               ELSIF (#statCountChannelPos = #CONST_CHANNEL_POS1)
               THEN
                   #statCurrentPos2 := #statCountChannelPos;
                   #statTimeImpulseSave2 := #statDeltaTimeImpulse;
                   #statTimePauseSave2 := #statDeltaTimePause;
                   #statTimeToImpulse := #statTimeToImpulse + #statDeltaTimeImpulse + #statDeltaTimePause;

                   IF ((#statDeltaTimePause >= #TIME_PAUSE1_MIN)
                       AND (#statDeltaTimePause <= #TIME_PAUSE1_MAX))
                   THEN
                       #statChannelActive2 := true;
                       #statCountChannelPos := #CONST_CHANNEL_POS2; // go to next pos 2
                   END_IF;

                   IF ((#statDeltaTimePause >= #TIME_PAUSE2_MIN)
                       AND (#statDeltaTimePause <= #TIME_PAUSE2_MAX))
                   THEN
                       #statChannelActive2 := false;
                       #statChannelActive3 := true;
                       #statCountChannelPos := #CONST_CHANNEL_POS2; // go to next Pos 2
                   END_IF;

                   IF ((#statDeltaTimePause >= #TIME_PAUSE3_MIN)
                       AND (#statDeltaTimePause <= #TIME_PAUSE3_MAX))
                   THEN
                       #statChannelActive2 := false;
                       #statChannelActive3 := false;
                       #statChannelActive4 := true;
                       #statCountChannelPos := #CONST_INT_0;
                   END_IF;

               ELSIF (#statCountChannelPos = #CONST_CHANNEL_POS2)
               THEN
                   #statCurrentPos3 := #statCountChannelPos;
                   #statTimeImpulseSave3 := #statDeltaTimeImpulse;
                   #statTimePauseSave3 := #statDeltaTimePause;
                   #statTimeToImpulse := #statTimeToImpulse + #statDeltaTimeImpulse + #statDeltaTimePause;

                   IF ((#statDeltaTimePause >= #TIME_PAUSE1_MIN)
                       AND (#statDeltaTimePause <= #TIME_PAUSE1_MAX))
                   THEN
                       #statChannelActive3 := true;
                       #statCountChannelPos := #CONST_CHANNEL_POS3; // go to next pos 3
                   END_IF;

                   IF ((#statDeltaTimePause >= #TIME_PAUSE2_MIN)
                       AND (#statDeltaTimePause <= #TIME_PAUSE2_MAX))
                   THEN
                       #statChannelActive3 := false;
                       #statChannelActive4 := true;
                       #statCountChannelPos := #CONST_INT_0;
                   END_IF;

               ELSIF (#statCountChannelPos = #CONST_CHANNEL_POS3)
               THEN
                   #statCurrentPos4 := #statCountChannelPos;
                   #statTimeImpulseSave4 := #statDeltaTimeImpulse;
                   #statTimePauseSave4 := #statDeltaTimePause;
                   #statTimeToImpulse := #statTimeToImpulse + #statDeltaTimeImpulse + #statDeltaTimePause;

                   IF ((#statDeltaTimePause >= #TIME_PAUSE1_MIN)
                       AND (#statDeltaTimePause <= #TIME_PAUSE1_MAX))
                   THEN
                       #statChannelActive4 := true;
                   END_IF;
                   #statCountChannelPos := #CONST_INT_0; // go to pos 0
               END_IF;
           END_IF;

       #STATE_ERROR:
           #error := true;
           #busy := false;
           #done := false;
           #statSysTimerStart := false;
           #statWatchDogTimerRisingStart := false;
           #statWatchDogTimerFallingStart := false;
           #status := #statStatus;
           #statStatus := #CONST_WORD_0;
           #statIndex := #STATE_IDLE;
       ELSE
           #statIndex := #STATE_IDLE;
   END_CASE;

   #instWatchDogTimerRising(IN := #statWatchDogTimerRisingStart,
                      PT := #CONST_WATCHDOG_TIMER,
                      Q=>#statWatchDogTimerRisingStop,
                      ET=>#statWatchDogTimerRisingRun);

   #instWatchDogTimerFalling(IN:=#statWatchDogTimerFallingStart,
                             PT:=#CONST_WATCHDOG_TIMER,
                             Q=>#statWatchDogTimerFallingStop,
                             ET=>#statWatchDogTimerFallingRun);


   #instSysTimer(IN:=#statSysTimerStart,
                 PT:=#CONST_CYCLETIME_TIMER,
                 Q=>#statSysTimerStop,
                 ET=>#statSysTimerRun);

   IF (#statWatchDogTimerRisingStop = TRUE)
       OR (#statWatchDogTimerFallingStop =true)
   THEN
       #statIndex := #STATE_ERROR;
       #statStatus := #CONST_ERROR_WATCHDOG_TIMER;
   END_IF;


   IF (#statSysTimerStop=true)
   THEN
       #statIndex := #STATE_ERROR;
       #statStatus := #CONST_ERROR_CYCLETIME_TIMER;
   END_IF;

   //Edge control
   #statImpulseOld := #impulse;
   #statResetOld := #reset;

   // Cycle time control
   #statSysTimeOld := #statSysTime;
END_FUNCTION_BLOCK

// ===== library types =====

TYPE "M_ZLT"
VERSION : 0.1
   STRUCT
      Fehl_empf : Bool;
      Fehl_Krit : Bool;
      Fehl_TO : Bool;
      STue_Abgl : Bool;
      Mel_Überlauf : Bool;
      Mel_Parameter : Bool;
      F_PW_Nr : Bool;
      Fehl_Senden : Bool;
      RM_ArbZeit : Bool;
      RM_Pause : Bool;
      RM_Schicht_1 : Bool;
      RM_Schicht_2 : Bool;
      RM_Schicht_3 : Bool;
      RM_Schicht_4 : Bool;
      RM_LSp : Bool;
      RM_Res : Bool;
   END_STRUCT;
END_TYPE

// folder: Audi_Bib/GF_Bausteine

FUNCTION_BLOCK "GF_GrFunktionen"   // FB200, SCL
{ S7_Optimized_Access := 'TRUE' }
VERSION : 0.1
   VAR_INPUT
      Quit_F : Bool;   // Quittierung Sicherheit/ Wiedereingliederung
      Init : Bool;
      TW_Res : Time;   // Zeitwert Resetzeit in 0,1s max 25sec
      TW_FQuit : Time;
   END_VAR
   VAR_OUTPUT
      F_Quit : Bool;
   END_VAR
   VAR
      R_TRIG_Instance : R_TRIG;
   END_VAR
   VAR RETAIN
      HMAnlauf : Bool;   // Hilfsmerker Anlauf
      HMAnl_ab : Bool;
      A_F_Quit : Bool;
      Quit_F_ab : Bool;
      Anl_Verzögerung : TON_TIME;
      IEC_Timer_0_Instance : TOF_TIME;
      Ret_SNC_RTCB : Int;
      Ret_WR_SYS : Int;
      T_Start_1 : Bool;
      T_abgel_1 : Bool;
      T_Start_2 : Bool;
      T_abgel_2 : Bool;
      Lfd_Nr_HText_1 : Int;
      Lfd_Nr_HText_2 : Int;
      "Tverz_Info-Text_1" : TON_TIME;
      "TVerz_Info-Text_2" : TON_TIME;
   END_VAR
   VAR_TEMP
      Stell_Zeit : DTL;
      S_1 : String;
      Ret_VAl : Int;
      T_Int : Int;
      UInt_1 : UInt;
      Zeit : String;
      Datum : String;
      X_Anzahl : Int;
      x : Int;
      Dat_Uhrz : String[24];
      HStr_3 : String[3];
   END_VAR
BEGIN
   (* Funktionsbeschreibung:                                                   Stand 6.5.2015
   ----------------------


   Baustein-Änderungen:
   --------------------
   Stand 9.6.2011  Identisch mit FB60 V 1.9 NSU Stand 18.2.2011
   Stand 22.9.2011  CPU-Meldungen aus Fehlermelde-OB´s angepasst (Adresse)
                    gemessene Zykluszeit "Mit" Rücksetzung eingefügt
   Stand 6.5.2015   Umstellung Takt-Merker auf Cyclic Interrupt-OB_s dadurch werden
                    keine CPU-Taktmerker mehr benötigt
   V0.1.7    Remanenz und Speicherreserve für Laden eingestellt



   *)                

   "VKE0":= false; "VS".VKE0 := false;                               // Vorbesetzung Systemmerker
   "VKE1":= true; "VS".VKE1 := true;
   "VS".Null := false;
   "VS".Eins := TRUE;
   "VS".Ohne := false;
   "VS".Mit := true;
   "VS".Mel_int := false;
   "VS".Kon_int := false;
   "VS".Sifa_int := false;

   "VS".Steu_ein := True;

   "VS".BliL := "VS"."Takt_0,5s";            // Blinktakte 500mSek
   "VS".BliS := "VS"."Takt_0,2s";              // Blinktakt 250mSek

   "VS"."ZTakt_0,1s" := false;                 // Zähltakt 100mSek.
   IF "VS"."Trig_0,1s" THEN
      "VS"."ZTakt_0,1s" := true;
      "VS"."Trig_0,1s" := false;
   END_IF;
   #R_TRIG_Instance(CLK:="VS"."Takt_0,5s", Q=>"VS".ZTakt_1s);               // Zähltakt 1Sekunde


   IF #HMAnlauf THEN #HMAnlauf:= false; "VS".Neustart:= false;  END_IF;       // Anlauf nach Neustart
   IF "VS".Neustart  THEN "VS".Anl_Verlae:= true; #HMAnlauf:= true; END_IF;
   #Anl_Verzögerung(IN:="VS".Anl_Verlae, PT:=#TW_Res,Q=>#HMAnl_ab );
   IF #HMAnl_ab THEN "VS".Anl_Verlae:= false; END_IF;
   "VS".Reset := "VS".Anl_Verlae;

   IF #HMAnl_ab OR "VS".Neustart  THEN #A_F_Quit:= true; END_IF;                        // F-Quit bilden
   #IEC_Timer_0_Instance(IN:=#A_F_Quit,  PT:=#TW_FQuit, Q=>#Quit_F_ab);
   IF #Quit_F_ab THEN #A_F_Quit:= false; END_IF;
   #F_Quit:= #A_F_Quit;

   // ************* Zykluszeit
   "GF_Zeitmessung"(Reset:="GF_Grund_DB".Res_Zeit[1],    // Zykluszeit errechnen
                    Mes_auswert:=true,
                    Zeit:="GF_Grund_DB".Zeit[1]);


   // CPU Zeit Stellen  Anstoss von Panel oder aus ZLT-Paket(Zeit-Synchronisation)
   IF "GF_Grund_DB".Stellbits.OP_Stell OR "GF_Grund_DB".Stellbits.Stell_ASCII THEN
      IF "GF_Grund_DB".Stellbits.Stell_ASCII THEN                                          // Zeitsynchronisation
         "GF_Grund_DB".Stellbits.Stell_ASCII := FALSE;                                                           //Stellzeit Typ DTL aus ASCII bilden
         Chars_TO_Strg(Chars := "GF_Grund_DB".Stell_Datum_Uhrzeit_ASCI.Jahr, pChars := 0, Cnt := 4,  Strg => #S_1);      //    Jahr
         #Stell_Zeit.YEAR := S_CONV(#S_1);
         Chars_TO_Strg(Chars := "GF_Grund_DB".Stell_Datum_Uhrzeit_ASCI.Monat, pChars := 0, Cnt := 2, Strg => #S_1);      //    Monat
         #Stell_Zeit.MONTH := S_CONV(#S_1);
         Chars_TO_Strg(Chars := "GF_Grund_DB".Stell_Datum_Uhrzeit_ASCI.Tag, pChars := 0, Cnt := 2, Strg => #S_1);        //    Tag
         #Stell_Zeit.DAY := S_CONV(#S_1);

         Chars_TO_Strg(Chars := "GF_Grund_DB".Stell_Datum_Uhrzeit_ASCI.Stunde, pChars := 0, Cnt := 2, Strg => #S_1);     //    Stunde
         #Stell_Zeit.HOUR := S_CONV(#S_1);
         Chars_TO_Strg(Chars := "GF_Grund_DB".Stell_Datum_Uhrzeit_ASCI.Minute, pChars := 0, Cnt := 2, Strg => #S_1);     //    Minute
         #Stell_Zeit.MINUTE := S_CONV(#S_1);
         Chars_TO_Strg(Chars := "GF_Grund_DB".Stell_Datum_Uhrzeit_ASCI.Sekunde, pChars := 0, Cnt := 2, Strg => #S_1);    //    Sekunde
         #Stell_Zeit.SECOND := S_CONV(#S_1);

         Chars_TO_Strg(Chars := "GF_Grund_DB".Stell_Datum_Uhrzeit_ASCI.MilliSek, pChars := 0, Cnt := 3, Strg => #S_1);   //    Millisekunde
         #Stell_Zeit.NANOSECOND := S_CONV(#S_1);
         #S_1 := S_CONV("GF_Grund_DB".Stell_Datum_Uhrzeit_ASCI.Wochentag);                                       //    Wochentag
         #Stell_Zeit.WEEKDAY := S_CONV(#S_1);

         "GF_Grund_DB".Stell_Datum_Uhrzeit := #Stell_Zeit;
         END_IF;

      IF "GF_Grund_DB".Stellbits.OP_Stell THEN                                 // Uhrzeit stellen von TP (Format DTL)
         "GF_Grund_DB".Stellbits.OP_Stell := false;
         #Stell_Zeit := "GF_Grund_DB".Stell_Datum_Uhrzeit;
      END_IF;

      #Ret_WR_SYS := WR_SYS_T(#Stell_Zeit);           // Uhrzeit stellen
      "GF_Grund_DB".Ret_Val := #Ret_VAl;

      #Ret_SNC_RTCB := SNC_RTCB();                      // Zeitsynchronisation nachtriggern
   END_IF;
   #T_Int := #Ret_SNC_RTCB; #T_Int := #Ret_WR_SYS;


   // ******************* CPU-Zeit auslesen
   //  Datum
   #Ret_VAl:=RD_LOC_T("GF_Grund_DB".Akt_Datum_Uhrzeit);                                                           // Aktuelle Datum/Zeit im Format DTL
   #S_1:=S_CONV("GF_Grund_DB".Akt_Datum_Uhrzeit.YEAR);                                                      // Umsetzung DTL in ASCII  Jahr
   #S_1:=RIGHT(IN:=#S_1, L:=4);
   #UInt_1 := 4;
   Strg_TO_Chars(Strg:=#S_1, pChars:=0,Cnt=>#UInt_1 , Chars:="GF_Grund_DB".Akt_Datum_Uhrzeit_ASCII.Datum.Jahr);
   #Datum := #S_1;
   #S_1:=S_CONV("GF_Grund_DB".Akt_Datum_Uhrzeit.MONTH);                                                     // Monat 
   #S_1 := REPLACE(IN1 := #S_1, IN2 := '0', L := 1, P := 1);
   #S_1:=RIGHT(IN:=#S_1, L:=2);
   Strg_TO_Chars(Strg:=#S_1, pChars:=0,Cnt=>#UInt_1, Chars:="GF_Grund_DB".Akt_Datum_Uhrzeit_ASCII.Datum.Monat);
   #Datum :=CONCAT(IN1:=#Datum, IN2:=#S_1);
   #S_1:=S_CONV("GF_Grund_DB".Akt_Datum_Uhrzeit.DAY);                                                       // Tag
   #S_1 := REPLACE(IN1 := #S_1, IN2 := '0', L := 1, P := 1);
   #S_1 := RIGHT(IN := #S_1, L := 2);
   Strg_TO_Chars(Strg:=#S_1, pChars:=0,Cnt=>#UInt_1, Chars:="GF_Grund_DB".Akt_Datum_Uhrzeit_ASCII.Datum.Tag);
   "GF_Grund_DB".Akt_Datum_Uhrzeit_ASCII.Datum.YYYYMMDD := CONCAT(IN1 := #Datum, IN2 := #S_1);

   // ***************** Zeit
   #S_1:=S_CONV("GF_Grund_DB".Akt_Datum_Uhrzeit.HOUR);                                                       // Stunde
   #S_1 := REPLACE(IN1 := #S_1, IN2 := '0', L := 1, P := 1);
   #S_1 := RIGHT(IN := #S_1, L := 2);
   Strg_TO_Chars(Strg:=#S_1, pChars:=0,Cnt=>#UInt_1, Chars:="GF_Grund_DB".Akt_Datum_Uhrzeit_ASCII.Zeit.Stunde);
   #Zeit := #S_1;
   #S_1:=S_CONV("GF_Grund_DB".Akt_Datum_Uhrzeit.MINUTE);                                                    // Minute
   #S_1 := REPLACE(IN1 := #S_1, IN2 := '0', L := 1, P := 1);
   #S_1:=RIGHT(IN:=#S_1, L:=2);
   Strg_TO_Chars(Strg:=#S_1, pChars:=0,Cnt=>#UInt_1, Chars:="GF_Grund_DB".Akt_Datum_Uhrzeit_ASCII.Zeit.Minute);
   #Zeit := CONCAT(IN1 := #Zeit, IN2 := #S_1); 
   #S_1:=S_CONV("GF_Grund_DB".Akt_Datum_Uhrzeit.SECOND);                                                    // Sekunde
   #S_1 := REPLACE(IN1 := #S_1, IN2 := '0', L := 1, P := 1);
   #S_1:=RIGHT(IN:=#S_1, L:=2);
   Strg_TO_Chars(Strg:=#S_1, pChars:=0,Cnt=>#UInt_1, Chars:="GF_Grund_DB".Akt_Datum_Uhrzeit_ASCII.Zeit.Sekunde);
   "GF_Grund_DB".Akt_Datum_Uhrzeit_ASCII.Zeit.HHMMSS := CONCAT(IN1 := #Zeit, IN2 := #S_1);

   #S_1:=S_CONV("GF_Grund_DB".Akt_Datum_Uhrzeit.NANOSECOND);                                                                                                                        
   // Milli-Sekunde
   #S_1:=MID(IN:=#S_1, L:=3, P:=3);
   Strg_TO_Chars(Strg:=#S_1, pChars:=0,Cnt=>#UInt_1, Chars:="GF_Grund_DB".Akt_Datum_Uhrzeit_ASCII.Zeit.MilliSek);
   #S_1:=S_CONV("GF_Grund_DB".Akt_Datum_Uhrzeit.WEEKDAY);                                                   // Wochentag
   #S_1:=RIGHT(IN:=#S_1, L:=1);
   "GF_Grund_DB".Akt_Datum_Uhrzeit_ASCII.Wochentag :=S_CONV(#S_1);

   //*********** Zeitformat für MA-PC (Fuchs-Paket) bereitstellen
   #Dat_Uhrz := "GF_Grund_DB".Akt_Datum_Uhrzeit_ASCII.Datum.YYYYMMDD;
   #Dat_Uhrz := INSERT(IN1 := #Dat_Uhrz, IN2 := '-', P := 4);                                          // YYYY-MMTT
   #Dat_Uhrz := INSERT(IN1 := #Dat_Uhrz, IN2 := '-', P := 7);                                          // YYYY-MM-TT
   #Dat_Uhrz := INSERT(IN1 := #Dat_Uhrz, IN2 := '  ', P := 11);                                        // YYYY-MM-TT__
   #Dat_Uhrz := INSERT(IN1 := #Dat_Uhrz, IN2 := "GF_Grund_DB".Akt_Datum_Uhrzeit_ASCII.Zeit.HHMMSS, P := 12);   // 
   #Dat_Uhrz := INSERT(IN1 := #Dat_Uhrz, IN2 := ':', P := 14);                                         // YYYY-MM-TT__hh:mmss
   #Dat_Uhrz := INSERT(IN1 := #Dat_Uhrz, IN2 := ':', P := 17);                                         // YYYY-MM-TT__hh:mm:ss
   #Dat_Uhrz := INSERT(IN1 := #Dat_Uhrz, IN2 := ':', P := 20);                                         // YYYY-MM-TT__hh:mm:ss:
   Chars_TO_Strg(Chars := "GF_Grund_DB".Akt_Datum_Uhrzeit_ASCII.Zeit.MilliSek,
                 pChars := 0, Cnt := 3,Strg => #HStr_3);
   #Dat_Uhrz := INSERT(IN1 := #Dat_Uhrz, IN2 := #HStr_3, P := 21);                                     // YYYY-MM-TT__hh:mm:ss:mmm
   "GF_Grund_DB".Zeit_Ma_PC := #Dat_Uhrz;

   // *********  globale Visu Info-Texte nach 5 Sek freigaben
   IF "GF_Visu_allg".H_Text_1."umlfd.Nr" <> #Lfd_Nr_HText_1 AND "GF_Visu_allg".H_Text_1.Pult <> 'X'  THEN
      #Lfd_Nr_HText_1 := "GF_Visu_allg".H_Text_1."umlfd.Nr";
      #T_Start_1 := true;
   END_IF;
   #"Tverz_Info-Text_1"(IN := #T_Start_1, PT := T#5s, Q => #T_abgel_1);
   IF #T_abgel_1 THEN
      "GF_Visu_allg".H_Text_1."umlfd.Nr" := 0;
      "GF_Visu_allg".H_Text_1.Pult := 'X';
      "GF_Visu_allg".H_Text_1.Stellglied := ' ';
      "GF_Visu_allg".H_Text_1.H_Text := ' ';
      #T_Start_1 := false;
   END_IF;

   IF "GF_Visu_allg".H_Text_2."umlfd.Nr" <> #Lfd_Nr_HText_2 AND "GF_Visu_allg".H_Text_2.Pult <> 'X' THEN
      #Lfd_Nr_HText_2 := "GF_Visu_allg".H_Text_2."umlfd.Nr";
      #T_Start_2 := true;
   END_IF;
   #"TVerz_Info-Text_2"(IN := #T_Start_2, PT := T#5s, Q => #T_abgel_2);
   IF #T_abgel_2 THEN
      "GF_Visu_allg".H_Text_2."umlfd.Nr" := 0;
      "GF_Visu_allg".H_Text_2.Pult := 'X';
      "GF_Visu_allg".H_Text_2.Stellglied := ' ';
      "GF_Visu_allg".H_Text_2.H_Text := ' ';
      #T_Start_2 := false;
   END_IF;

   // ***********************  Initialisierungen
   IF #Init OR "VS".Neustart THEN
      #T_Start_1 := false;   #T_abgel_1 := false;
      #T_Start_2 := false;   #T_abgel_2 := false;

      "GF_Visu_allg".H_Text_1.Pult := 'X';
      "GF_Visu_allg".H_Text_1."umlfd.Nr" := 0;
      "GF_Visu_allg".H_Text_2.Pult := 'X';
      "GF_Visu_allg".H_Text_2."umlfd.Nr" := 0;

       #X_Anzahl := "GF_An_Vor_St".max_Anzahl;                         // An/Vorwahlen
       FOR #x := 1 TO #X_Anzahl DO                                     //   Eintrag Array-NR. in Array-Element NR
           "GF_An_Vor_St".An_Vorw[#x].AnVisu.Nr := #x;
           "GF_An_Vor_St".An_Vorw[#x].AnVisu.Bed_Station := 'xxxx';
           "GF_An_Vor_St".An_Vorw[#x].AnVisu.Bezeichnung := '    ';
           "GF_An_Vor_St".An_Vorw[#x].AnVisu.Status := 0;
       END_FOR;

       #X_Anzahl := "GF_LastSp_St".max_Anzahl;                         // Lastspannungen
       FOR #x := 1 TO #X_Anzahl DO                                     // Eintrag Array-NR. in Array-Element NR
           "GF_LastSp_St".LastSp[#x].AnVisu.Nr := #x;
           "GF_LastSp_St".LastSp[#x].AnVisu.Bed_Station := 'xxxx';
           "GF_LastSp_St".LastSp[#x].AnVisu.Bezeichnung := '    ';
           "GF_LastSp_St".LastSp[#x].AnVisu.Status := 0;
       END_FOR;

       #X_Anzahl := "GF_BetrArt_St".max_Anzahl;                        // Betriebsarten
       FOR #x := 1 TO #X_Anzahl DO                                     // Eintrag Array-NR. in Array-Element NR
           "GF_BetrArt_St".BetrArt[#x].AnVisu.Nr := #x;
           "GF_BetrArt_St".BetrArt[#x].AnVisu.Bed_Station := 'xxxx';
           "GF_BetrArt_St".BetrArt[#x].AnVisu.Bezeichnung := '    ';
           "GF_BetrArt_St".BetrArt[#x].AnVisu.Status := 0;
       END_FOR;

       #X_Anzahl := "GF_HBed_Obj_St".max_Anzahl;                       // Hand-Bedien-Objekte
       FOR #x := 1 TO #X_Anzahl DO                                     // Eintrag Array-NR. in Array-Element NR
           "GF_HBed_Obj_St".Modul[#x].Nr := #x;
       END_FOR;

       #X_Anzahl := 8;                                                 // Meldekanäle initialisieren
       FOR #x := 1 TO #X_Anzahl DO                                 
           "GF_Visu_allg".SS.Kanal[#x].Belegung.Pult_Name := 'xxxx';
       END_FOR;
   END_IF;
END_FUNCTION_BLOCK

FUNCTION "GF_Zeitmessung" : Void   // FC205, SCL
{ S7_Optimized_Access := 'TRUE' }
VERSION : 0.1
   VAR_INPUT
      Reset : Bool;   // Reset gemessene Zeiten
      Mes_auswert : Bool;   // 0 = Messung starten, 1 = Messung auswerten
   END_VAR
   VAR_IN_OUT
      Zeit : "GF_Zeit_Messung";
   END_VAR
   VAR_TEMP
      H_zeit : LReal;
   END_VAR
BEGIN
   (*
   aktuelle Baustein-Version 0.2.0

   User-Dokumentation über Shift F1
   Ablage im Projekt-Ordner Bereich UserDocumentation
   Doku-Datum 15.4.15

   Baustein-Historie ***********************************
   Version     Änderung
    0.2.x      Basis-Version


   *)


   IF #Reset OR "VS".Reset THEN                                          // gemessene Zeiten löschen
       #Zeit.akt := 0;
       #Zeit.min := 0;
       #Zeit.max := 0;
   END_IF;

   #H_zeit := RUNTIME(#Zeit.Speicher);                                  // aktuelle Zeit auslesen
   IF #Mes_auswert  THEN
      #H_zeit := #H_zeit * 1000000;
      #Zeit.akt := LREAL_TO_INT(#H_zeit);                               // umsetzen in INT
       IF #Reset OR "VS".Reset THEN
           #Zeit.max := #Zeit.akt;
           #Zeit.min := #Zeit.akt;
        ELSE
           IF #Zeit.akt > #Zeit.max THEN
               #Zeit.max := #Zeit.akt;
           END_IF;
           IF #Zeit.akt < #Zeit.min THEN
               #Zeit.min := #Zeit.akt;
            END_IF;
        END_IF;
   END_IF;
END_FUNCTION

// ===== library: CodeBlockByCopyVersionObject "None" =====

// ===== library: CodeBlockByCopyVersionObject "None" =====

// ===== library: UserTypeByCopyVersionObject "None" =====

// ===== library: UserTypeByCopyVersionObject "None" =====

// ===== library: UserTypeByCopyVersionObject "None" =====

// ===== library: CodeBlockByCopyVersionObject "None" =====

(* ===== HMI "HMI_RT_1" =====

ScreenModuleEditorView "typeSlot" 640x480
   Rectangle "Rectangle_2" at 18,19 size 49x139
      Visibility <- "SlotUsed"
      Appearance <- "SlotErrorState"
   TextField "Text field_5" at 18,23 size 49x25; Text '00'
      Visibility <- "SlotUsed"
*)

(* ===== HMI "HMI_RT_1" =====

ScreenModuleEditorView "typeDevice" 640x480
   Button "Schaltfläche_3" at 90,10 size 110x110; TextOff 'Text'
      Visibility <- "DeviceNumber"
   Rectangle "Rectangle_1" at 90,10 size 110x110
      Visibility <- "DeviceNumber"
      Appearance <- "ErrorState"
   IOField "EA-Feld_1" at 90,10 size 110x110; FormatPattern 999
      Visibility <- "DeviceNumber"
      ProcessValue <- "DeviceNumber"
*)

(* ===== HMI "HMI_RT_1" =====
system functions are stored by id; their names below are inferred from use

HMI tags "Standard-Variablentabelle"
   "showValues" : Bool, internal

ScreenModuleEditorView "SDC_EMS_TS_klein_unten_movLi" 1024x768
   Group "Group" at 78,28 size 49x65
      HorizontalMovement <- "EMS_SEK.DRIVE_POS_%"
   IOField "Hoist_Pos_moving" at 84,78 size 38x12; FormatPattern 9999
      Appearance <- "EMS_SEK.STAT_1"
      ProcessValue <- "EMS_SEK.HOIST_POS"
      Visibility <- "showValues"
   IOField "Drive_Pos_moving" at 78,67 size 49x12; FormatPattern 9999999
      Appearance <- "EMS_SEK.STAT_1"
      ProcessValue <- "EMS_SEK.DRIVE_POS"
      Visibility <- "showValues"
   IOField "EMS_Nr" at 81,48 size 43x20; FormatPattern 999
      Visibility <- "EMS_SEK.EMS_ID"
      ProcessValue <- "EMS_SEK.EMS_ID"
      Appearance <- "EMS_SEK.STAT_1"
   IOField "ERROR_No" at 81,29 size 43x20; FormatPattern 999
      Appearance <- "EMS_SEK.ERROR"
      ProcessValue <- "EMS_SEK.ERROR"
      Visibility <- "EMS_SEK.ERROR"
   Button "S_EMS_Nr_uebergeben" at 81,29 size 43x53; TextOff 'Text'
      on Click: "Uebergabe_EMS_Nr"(); InvertBit("open_EMS_STAT")
      ObjectEnable <- "EMS_SEK.EMS_ID"
      Visibility <- "EMS_SEK.EMS_ID"

VB script "Uebergabe_EMS_Nr"
   ' EMS- Nummer übergeben
   
   ' Groiß Andreas 
   ' Siemens AG Österreich 
   ' Linz Kraußstraße 1-7 
   ' I IA AS SO AP2 Surface Technology & Assembly
   ' 12.09.2012 
   
   	If SmartTags("EMS_SEK.EMS_ID") > 0 Then
   	
   		SmartTags("EMS_Nr") = SmartTags("EMS_SEK.EMS_ID")
   		
   	Else
   		
   		SmartTags("EMS_Nr") = 1
   		
   	End If

VB script "showValues"
   'Tip:
   ' 1. Verwenden Sie die Tastenkombination <CTRL+SPACE> oder <CTRL+I>, um eine Liste aller Objekte und Funktionen zu öffnen
   ' 2. Schreiben Sie den Code unter Verwendung des HMI Runtime Objekts.
   '  Beispiel: HmiRuntime.Screens("Screen_1").
   ' 3. Verwenden Sie die Tastenkombination <CTRL+J>, um eine Objektreferenz zu erstellen.
   'Schreiben Sie den Code ab dieser Position:
   If SmartTags("EMS_SEK.EMS_ID")>0 And SmartTags("Pos_sichtbar") Then
   	SmartTags("showValues") = True
   Else
   	SmartTags("showValues") = False
   End If
*)

(* ===== HMI "HMI_RT_2" =====
system functions are stored by id; their names below are inferred from use
connection "SDC_PLC": ETHERNET, S7_1500_OMS

HMI tags "Standard-Variablentabelle"
   "Trigger" : Int, internal
   "TP_Online" : Int, internal
   "_BildNr_aktuell" : Int, internal
   "__Pult_Name" : Int, internal
   "__Pult_Name(1)" : WString[10], internal
   "test" : Int, internal
   "LinePLC1_RD_ready" : Bool = PLC LinePLC1_RD_ready AT %I4248.0, 1 s
   "DiagStatusUpdate" : Bool = PLC DiagStatusUpdate AT %M1.1, 1 s
   "EMS_Carrier_Spacing" : Int = PLC EMS.Carrier_Spacing, 1 s
   "EMS_Coarse_Decel_Speed" : Word = PLC EMS.CoarseDecelSpeed AT %DB1.DBW0, 1 s
   "EMS_Coarse_Position_Decel_Offset" : Word = PLC EMS.CoarsePositionDecelOffset AT %DB1.DBW0, 1 s
   "EMS_Coarse_Position_Tolerance" : Word = PLC EMS.CoarsePositionTolerance AT %DB1.DBW0, 1 s
   "EMS_Fine_Decel_Speed" : Word = PLC EMS.FineDecelSpeed AT %DB1.DBW0, 1 s
   "EMS_Fine_Posistion_Tolerance" : Word = PLC EMS.FinePositionTolerance AT %DB1.DBW0, 1 s
   "EMS_Fine_Position_Decel_Offset" : Word = PLC EMS.FinePositionDecelOffset AT %DB1.DBW0, 1 s
   "EMS_Production_Spacing" : Word = PLC EMS.Production_Spacing, 1 s
   "EMS_Production_Zone_Speed" : Word = PLC EMS.ProductionZnSpeed AT %DB1.DBW0, 1 s
   "Temp_Placeholder" : Int = PLC Temp_Int AT %MW56, 1 s
   "CARRIER #01   CURRENT" : Int = PLC "CARRIER #01   CURRENT" AT %MW72, 1 s
   "CARRIER #01   G120D Status WORD.0(1)" : Bool = PLC "CARRIER #01   G120D STATUS WORD.0" AT %M76.0, 1 s
   "CARRIER #01   G120D Status WORD.1(1)" : Bool = PLC "CARRIER #01   G120D STATUS WORD.1" AT %M76.1, 1 s
   "CARRIER #01   G120D Status WORD.10(1)" : Bool = PLC "CARRIER #01   G120D STATUS WORD.10" AT %M77.2, 1 s
   "CARRIER #01   G120D Status WORD.11(1)" : Bool = PLC "CARRIER #01   G120D STATUS WORD.11" AT %M77.3, 1 s
   "CARRIER #01   G120D Status WORD.12(1)" : Bool = PLC "CARRIER #01   G120D STATUS WORD.12" AT %M77.4, 1 s
   "CARRIER #01   G120D Status WORD.13(1)" : Bool = PLC "CARRIER #01   G120D STATUS WORD.13" AT %M77.5, 1 s
   "CARRIER #01   G120D Status WORD.14(1)" : Bool = PLC "CARRIER #01   G120D STATUS WORD.14" AT %M77.6, 1 s
   "CARRIER #01   G120D Status WORD.15(1)" : Bool = PLC "CARRIER #01   G120D STATUS WORD.15" AT %M77.7, 1 s
   "CARRIER #01   G120D Status WORD.2(1)" : Bool = PLC "CARRIER #01   G120D STATUS WORD.2" AT %M76.2, 1 s
   "CARRIER #01   G120D Status WORD.3(1)" : Bool = PLC "CARRIER #01   G120D STATUS WORD.3" AT %M76.3, 1 s
   "CARRIER #01   G120D Status WORD.4(1)" : Bool = PLC "CARRIER #01   G120D STATUS WORD.4" AT %M76.4, 1 s
   "CARRIER #01   G120D Status WORD.5(1)" : Bool = PLC "CARRIER #01   G120D STATUS WORD.5" AT %M76.5, 1 s
   "CARRIER #01   G120D Status WORD.6(1)" : Bool = PLC "CARRIER #01   G120D STATUS WORD.6" AT %M76.6, 1 s
   "CARRIER #01   G120D Status WORD.7(1)" : Bool = PLC "CARRIER #01   G120D STATUS WORD.7" AT %M76.7, 1 s
   "CARRIER #01   G120D Status WORD.8(1)" : Bool = PLC "CARRIER #01   G120D STATUS WORD.8" AT %M77.0, 1 s
   "CARRIER #01   G120D Status WORD.9(1)" : Bool = PLC "CARRIER #01   G120D STATUS WORD.9" AT %M77.1, 1 s
   "CARRIER #01   G120D STATUS WORD.0" : Bool = PLC "CARRIER #01   G120D STATUS WORD.0" AT %M76.0, 1 s
   "CARRIER #01   G120D STATUS WORD.1" : Bool = PLC "CARRIER #01   G120D STATUS WORD.1" AT %M76.1, 1 s
   "CARRIER #01   G120D STATUS WORD.10" : Bool = PLC "CARRIER #01   G120D STATUS WORD.10" AT %M77.2, 1 s
   "CARRIER #01   G120D STATUS WORD.11" : Bool = PLC "CARRIER #01   G120D STATUS WORD.11" AT %M77.3, 1 s
   "CARRIER #01   G120D STATUS WORD.12" : Bool = PLC "CARRIER #01   G120D STATUS WORD.12" AT %M77.4, 1 s
   "CARRIER #01   G120D STATUS WORD.13" : Bool = PLC "CARRIER #01   G120D STATUS WORD.13" AT %M77.5, 1 s
   "CARRIER #01   G120D STATUS WORD.14" : Bool = PLC "CARRIER #01   G120D STATUS WORD.14" AT %M77.6, 1 s
   "CARRIER #01   G120D STATUS WORD.15" : Bool = PLC "CARRIER #01   G120D STATUS WORD.15" AT %M77.7, 1 s
   "CARRIER #01   G120D STATUS WORD.2" : Bool = PLC "CARRIER #01   G120D STATUS WORD.2" AT %M76.2, 1 s
   "CARRIER #01   G120D STATUS WORD.3" : Bool = PLC "CARRIER #01   G120D STATUS WORD.3" AT %M76.3, 1 s
   "CARRIER #01   G120D STATUS WORD.4" : Bool = PLC "CARRIER #01   G120D STATUS WORD.4" AT %M76.4, 1 s
   "CARRIER #01   G120D STATUS WORD.5" : Bool = PLC "CARRIER #01   G120D STATUS WORD.5" AT %M76.5, 1 s
   "CARRIER #01   G120D STATUS WORD.6" : Bool = PLC "CARRIER #01   G120D STATUS WORD.6" AT %M76.6, 1 s
   "CARRIER #01   G120D STATUS WORD.7" : Bool = PLC "CARRIER #01   G120D STATUS WORD.7" AT %M76.7, 1 s
   "CARRIER #01   G120D STATUS WORD.8" : Bool = PLC "CARRIER #01   G120D STATUS WORD.8" AT %M77.0, 1 s
   "CARRIER #01   G120D STATUS WORD.9" : Bool = PLC "CARRIER #01   G120D STATUS WORD.9" AT %M77.1, 1 s
   "CARRIER #01   POSITION" : Int = PLC "CARRIER #01   POSITION" AT %MW78, 1 s
   "CARRIER #01 480VPowerOn_MDCB1" : Bool = PLC "CARRIER #01 480VPowerOn_MDCB1" AT %M80.0, 1 s
   "CARRIER #01 CrashDetectSW" : Bool = PLC "CARRIER #01 CrashDetectSW" AT %M80.1, 1 s
   "CARRIER #01 DCsupplyOnPSCB2" : Bool = PLC "CARRIER #01 DCsupplyOnPSCB2" AT %M80.2, 1 s
   "CARRIER #01 FaultLight_LH" : Bool = PLC "CARRIER #01 FaultLight_LH" AT %M80.3, 1 s
   "CARRIER #01 FaultLight_RH" : Bool = PLC "CARRIER #01 FaultLight_RH" AT %M80.4, 1 s
   "Carrier #01 HMI 1 Status0.5(1)" : Bool = PLC "CARRIER #01   1 STATUS [0].5" AT %M80.5, 1 s
   "CARRIER #01 PB1_ProdHoldLH" : Bool = PLC "CARRIER #01 PB1_ProdHoldLH" AT %M80.6, 1 s
   "CARRIER #01 PB2_ResetLH" : Bool = PLC "CARRIER #01 PB2_ResetLH" AT %M80.7, 1 s
   "CARRIER #01 PB3_ProdHoldRH" : Bool = PLC "CARRIER #01 PB3_ProdHoldRH" AT %M81.0, 1 s
   "CARRIER #01 PB4_ResetRH" : Bool = PLC "CARRIER #01 PB4_ResetRH" AT %M81.1, 1 s
   "CARRIER #01 RunLight_LH" : Bool = PLC "CARRIER #01 RunLight_LH" AT %M81.2, 1 s
   "CARRIER #01 RunLight_RH" : Bool = PLC "CARRIER #01 RunLight_RH" AT %M81.3, 1 s
   "CARRIER #01 SitopSelectStatus" : Bool = PLC "CARRIER #01 SitopSelectStatus" AT %M81.4, 1 s
   "CARRIER #01 SpareInput(2_1)" : Bool = PLC "CARRIER #01 SpareInput(2_1)" AT %M81.5, 1 s
   "CARRIER #01 SpareInput(2_2)" : Bool = PLC "CARRIER #01 SpareInput(2_2)" AT %M81.6, 1 s
   "CARRIER #01 SpareInput(2_3)" : Bool = PLC "CARRIER #01 SpareInput(2_3)" AT %M81.7, 1 s
   "CARRIER #01 SpareInput(2_4)" : Bool = PLC "CARRIER #01 SpareInput(2_4)" AT %M82.0, 1 s
   "CARRIER #01 SpareInput(2_5)" : Bool = PLC "CARRIER #01 SpareInput(2_5)" AT %M82.1, 1 s
   "CARRIER #01 SpareInput(2_6)" : Bool = PLC "CARRIER #01 SpareInput(2_6)" AT %M82.2, 1 s
   "CARRIER #01 SpareInput(2_7)" : Bool = PLC "CARRIER #01 SpareInput(2_7)" AT %M82.3, 1 s
   "CARRIER #01 SpareInput(4_1)" : Bool = PLC "CARRIER #01 SpareInput(4_1)" AT %M82.4, 1 s
   "CARRIER #01 SpareInput(4_14)" : Bool = PLC "CARRIER #01 SpareInput(4_14)" AT %M82.5, 1 s
   "CARRIER #01 SpareInput(4_15)" : Bool = PLC "CARRIER #01 SpareInput(4_15)" AT %M82.6, 1 s
   "CARRIER #01 SpareInput(4_16)" : Bool = PLC "CARRIER #01 SpareInput(4_16)" AT %M82.7, 1 s
   "CARRIER #01 SpareInput(4_17)" : Bool = PLC "CARRIER #01 SpareInput(4_17)" AT %M83.0, 1 s
   "CARRIER #01 SpareInput(4_2)" : Bool = PLC "CARRIER #01 SpareInput(4_2)" AT %M83.1, 1 s
   "CARRIER #01 SpareInput(4_5)" : Bool = PLC "CARRIER #01 SpareInput(4_5)" AT %M83.2, 1 s
   "CARRIER #01 SpareInput(4_6)" : Bool = PLC "CARRIER #01 SpareInput(4_6)" AT %M83.3, 1 s
   "CARRIER #01 SpareInput(4_7)" : Bool = PLC "CARRIER #01 SpareInput(4_7)" AT %M83.4, 1 s
   "CARRIER #01 SpareOutput(5_5)" : Bool = PLC "CARRIER #01 SpareOutput(5_5)" AT %M83.5, 1 s
   "CARRIER #01 SpareOutput(5_6)" : Bool = PLC "CARRIER #01 SpareOutput(5_6)" AT %M83.6, 1 s
   "CARRIER #01 SpareOutput(5_7)" : Bool = PLC "CARRIER #01 SpareOutput(5_7)" AT %M83.7, 1 s
   "CARRIER #01 SpareSafetyOutput(3_1)" : Bool = PLC "CARRIER #01 SpareSafetyOutput(3_1)" AT %M84.0, 1 s